// TIA Portal project "test_program" (V15)

(* hardware
DEVICE "S71500/ET200MP station_1"  S7-1500 station
   slot 0: "Rail_0"  Rack  6ES7 590-1***0-0AA0
   slot 0: "PM 70W 120/230VAC"  PM 70W 120/230VAC  6EP1332-4BA00
   slot 1: "PLC_1"  CPU 1511-1 PN  6ES7 511-1AK00-0AB0  V1.6
   slot 2: "DI 16x24VDC HF_1"  DI 16x24VDC HF  6ES7 521-1BH00-0AB0  V2.0
   slot 3: "DQ 16x24VDC/0.5A ST_1"  DQ 16x24VDC/0.5A ST  6ES7 522-1BH00-0AB0  V2.0
DEVICE "SCALANCE X005"  SCALANCE X-Station
   slot 0: "SCALANCE X rack"  Rail
   slot 0: "Switch_1"  6GK5 005-0BA00-1AA3  V1.0
DEVICE "GSD device_1"  GSD.Device.PN
   slot 0: "Rack"  Rack  V1.0
   slot 0: "INpactPIR"  Standard  INpact-PIR  V5.07
      slot 0: "Standard"  Standard
      slot 1: "Interface"  Interface
         slot 1: "Port 1"  Port 1
         slot 2: "Port 2"  Port 2
*)

// ===== PLC "PLC_1"  CPU 1511-1 PN =====
// protected blocks, not shown: "PDSql_1500_FB"

VAR_GLOBAL   // PLC tag table "Default tag table"
   "AlwaysTrue" AT %M0.1 : Bool;
   "AlwaysFalse" AT %M0.2 : Bool;
END_VAR

TYPE "part_processing_data"
   STRUCT
      sPartGroupID : String;
      rAFM_Param_1 : Real;
      rAFM_Param_2 : Real;
      rAFM_Param_3 : Real;
      sPartID_1 : String;
      iPartID_2 : UDInt;
   END_STRUCT;
END_TYPE

// folder: Data Types

TYPE "tConnection"
   STRUCT
      IP1 : USInt;
      IP2 : USInt;
      IP3 : USInt;
      IP4 : USInt;
      Port : UDInt;
      ConnID : Conn_Ouc;
      HW : Hw_Interface;
      Timeout : Time;
   END_STRUCT;
END_TYPE

TYPE "tSqlTable_1200"
   STRUCT
      ColumnCount : UInt;
      RowCount : UInt;
      MaxColumns : UInt := 10;
      MaxRows : UInt := 10;
      MaxStringLength : USInt := 50;
      Columns : Array[1..10] of "tColumn_1200";
   END_STRUCT;
END_TYPE

TYPE "tColumn_1200"
   STRUCT
      "Name" : String;   // Column name
      UserType : Byte;   // Unique generator of row
      "Type" : Byte;   // MSSQL-Data-Type of column
      LenSize : Byte;   // Number of bytes used for Length information of data
      TypeNumericPrecision : Byte;
      TypeNumericScale : Byte;
      Nullable : Bool;
      CaseSens : Bool;
      Identity : Bool;
      Computed : Bool;
      FixedLenCLRType : Bool;
      UsUpdatable : Byte;
      Rows : Array[1..10] of "tRow_1200";
   END_STRUCT;
END_TYPE

TYPE "tLicence"
   STRUCT
      LicKey1 : DWord;
      LicKey2 : DWord;
      LicKey3 : DWord;
      LicKey4 : DWord;
      LicKey5 : DWord;
   END_STRUCT;
END_TYPE

TYPE "tRow_1200"
   STRUCT
      "Bool" : Bool;
      Null : Bool;
      "DInt" : DInt;
      LReal : LReal;
      "String" : String[50];
      Datetime : DTL;
   END_STRUCT;
END_TYPE

TYPE "tSqlTable_1500"
   STRUCT
      ColumnCount : UInt;
      RowCount : UInt;
      MaxColumns : UInt := 10;
      MaxRows : UInt := 10;
      MaxStringLength : USInt := 50;
      Columns : Array[1..10] of "tColumn_1500";
   END_STRUCT;
END_TYPE

TYPE "tColumn_1500"
   STRUCT
      "Name" : String;   // Column name
      UserType : Byte;   // Unique generator of row
      "Type" : Byte;   // MSSQL-Data-Type of column
      LenSize : Byte;   // Number of bytes used for Length information of data
      TypeNumericPrecision : Byte;
      TypeNumericScale : Byte;
      Nullable : Bool;
      CaseSens : Bool;
      Identity : Bool;
      Computed : Bool;
      FixedLenCLRType : Bool;
      UsUpdatable : Byte;
      Rows : Array[1..10] of "tRow_1500";
   END_STRUCT;
END_TYPE

TYPE "tRow_1500"
   STRUCT
      "Bool" : Bool;
      Null : Bool;
      LInt : LInt;
      LReal : LReal;
      "String" : String[50];
      Datetime : DTL;
   END_STRUCT;
END_TYPE

TYPE "tLogin"
   STRUCT
      HostName : String[50];   // Hostname for database
      UserName : String[50];   // Username
      Password : String[50];   // Password
      Database : String[50];   // Database name
   END_STRUCT;
END_TYPE

TYPE "tQuery"
   STRUCT
      Query : Array[1..2] of String;
   END_STRUCT;
END_TYPE

TYPE "tCmd"
   STRUCT
      Connect : Bool;
      Disconnect : Bool;
      ExecuteQuery : Bool;
   END_STRUCT;
END_TYPE

TYPE "tStat"
   STRUCT
      Connected : Bool;
      Busy : Bool;
      ExecutedOK : Bool;
      Error : Bool;
      Status : Word;
      Message : String;
   END_STRUCT;
END_TYPE

// folder: 01_S7-1500

DATA_BLOCK "101_Simulation_IDB"   // DB1
{ S7_Optimized_Access := 'TRUE' }
VERSION : 0.1
// stored: InstanceOfName 101_Simulation
"101_Simulation"
BEGIN
END_DATA_BLOCK

DATA_BLOCK "InputsDB"   // DB2
{ S7_Optimized_Access := 'TRUE' }
VERSION : 0.1
   VAR
      part_processing_data : "part_processing_data";
   END_VAR
BEGIN
   part_processing_data.sPartGroupID := 'Deutz_ASML_10102A';
   part_processing_data.rAFM_Param_1 := 11.12;
   part_processing_data.rAFM_Param_2 := 4.98;
   part_processing_data.rAFM_Param_3 := 30.96;
   part_processing_data.sPartID_1 := 'ASML_JDK32_';
   part_processing_data.iPartID_2 := 100786;
END_DATA_BLOCK

DATA_BLOCK "DB_PDSql_1500"   // DB2010
{ S7_Optimized_Access := 'TRUE' }
VERSION : 0.1
   VAR
      Connection : "tConnection";
      Licence : "tLicence";
      Cmd : "tCmd";
      Stat : "tStat";
      Login : "tLogin";
      Query : "tQuery";
      SQLTable : "tSqlTable_1500";
   END_VAR
BEGIN
   Connection.IP1 := 192;
   Connection.IP2 := 168;
   Connection.IP3 := 2;
   Connection.IP4 := 1;
   Connection.Port := 1433;
   Login.Database := 'S7_1500_PLC';
   Login.Password := 'admin-6969';
   Login.UserName := 'sa';
   Login.HostName := 'EEEL1000332\SQLEXPRESS';
   Connection.ConnID := 1;
   Connection.HW := 64;
   Connection.Timeout := t#2s;
   Licence.LicKey1 := 16#67ABDCEB;
   Licence.LicKey2 := 16#28EC4AC9;
   Licence.LicKey3 := 16#D8D955FC;
   Licence.LicKey4 := 16#4A43863A;
   Licence.LicKey5 := 16#74F235FD;
END_DATA_BLOCK

// folder: 00_Functions

FUNCTION "LGF_Random_Real" : Real   // FC1, SCL
{ S7_Optimized_Access := 'TRUE' }
VERSION : 0.1
   VAR_OUTPUT
      error : Bool;
      status : Word;
      subfunctionStatus : Word;
   END_VAR
   VAR_TEMP
      tempTime : DTL;
      tempNanoSecondInDWord : DWord;
      tempTimeStatus : DWord;
      tempRandomValue : DWord;
   END_VAR
   VAR CONSTANT
      ZERO : Real;
      MAX_UDINT : UDInt := 4294967295;
      SUB_STATUS_NO_ERROR : Word := 16#0000;
      STATUS_FINISHED_NO_ERROR : Word := 16#0000;
      ERR_RD_SYS_T : Word := 16#8600;
   END_VAR
BEGIN
   REGION Block info header
       //=============================================================================
       // SIEMENS AG / (c)Copyright 2017
       //-----------------------------------------------------------------------------
       // Title:            LGF_Random_Real
       // Comment/Function: Generates a random real number between 0.0 and 1.0
       // Library/Family:   LGF(Library General Functions)
       // Author:           Siemens Digital Industry Support
       // Tested with:      S7-PLCSIM Advanced V2.0 SP1
       // Engineering:      TIA Portal V15 Update 2
       // Restrictions:     ENO disabled - error handling done by error and status
       // Requirements:     PLC (S7-1200 / S7-1500)
       //-------------------------------------------------------------------------------
       // Change log table:
       // Version  | Date       | Expert in charge       | Changes applied
       //----------|------------|------------------------|------------------------------
       // 01.00.00 27.01.2017  Siemens Industry Online Support
       //                      First released version
       // 01.00.01 17.08.2018  Siemens Industry Online Support
       //                      Upgrade: TIA V15 Update 2
       // 01.00.02 23.11.2018  Siemens Industry Online Support
       //                      Upgrade: TIA V15.1
       // 01.01.00 13.11.2019  Siemens Industry Presales Support
       //                      Renamed from "LGF_RandomBasic" to "LGF_Random_Real"
       //                      Regions, commens and costants are added
       // 03.00.00 23.04.2020  Siemens Industry Support
       //                      Set version to V3.0.0, harmonize the version of the whole library
       //=============================================================================
   END_REGION

   REGION Validation
       // Read system time
       #tempTimeStatus := INT_TO_WORD(RD_SYS_T(#tempTime));

       // Check return variable for error
       IF (#tempTimeStatus <> #SUB_STATUS_NO_ERROR) THEN
           #error := true;
           #status := #ERR_RD_SYS_T;
           #subfunctionStatus := #tempTimeStatus;
           #LGF_Random_Real := #ZERO;
           RETURN;
       END_IF;
   END_REGION

   REGION Calculating random number
       // Converting to double word so individual bytes can be addressed
       #tempNanoSecondInDWord := UDINT_TO_DWORD(#tempTime.NANOSECOND);

       // Calculate a random-start-value depending on the time
       #tempRandomValue.%B3 := #tempNanoSecondInDWord.%B0;
       #tempRandomValue.%B2 := #tempNanoSecondInDWord.%B1;
       #tempRandomValue.%B1 := #tempNanoSecondInDWord.%B2;
       #tempRandomValue.%B0 := #tempNanoSecondInDWord.%B3;

       // Norm the calculated random number: 0.0 <= Random_Real <= 1.0
       #LGF_Random_Real := UDINT_TO_REAL(DWORD_TO_UDINT(#tempRandomValue)) / UDINT_TO_REAL(#MAX_UDINT);

       #error := false;
       #status := #STATUS_FINISHED_NO_ERROR;
       #subfunctionStatus := #SUB_STATUS_NO_ERROR;
       // ENO mechanism is not used
       ENO := TRUE;
   END_REGION
END_FUNCTION

FUNCTION "fcRemovePlus" : String   // FC18, SCL
{ S7_Optimized_Access := 'TRUE' }
VERSION : 0.1
   VAR_INPUT
      STR : String;
   END_VAR
BEGIN
   //=============================================================================
   // PLCdirectSQL (c)Copyright 2019
   //-----------------------------------------------------------------------------
   // Library: fcRemovePlus
   // Tested with: S7-1200 FW 4.2 / S7-1500 FW 1.8
   // Engineering: TIA Portal 14
   // Requirements: S7-1200/1500
   // Functionality: Remove the first plus sign ("+") from a string
   //-----------------------------------------------------------------------------
   // Change log:
   // dd.mm.yyyy
   // 06.06.2019 Igor Filanda 1.0 First Release
   //=============================================================================

   IF FIND(IN1 := #STR, IN2 := '+') <> 0 THEN
       #fcRemovePlus := DELETE(IN := #STR, L := 1, P := FIND(IN1 := #STR, IN2 := '+'));
   ELSE
       #fcRemovePlus := #STR;
   END_IF;
END_FUNCTION

FUNCTION "fcDTLString" : String   // FC19, SCL
{ S7_Optimized_Access := 'TRUE' }
VERSION : 0.1
   VAR_INPUT
      dtlDatetime : DTL;
   END_VAR
   VAR_TEMP
      str : String;
   END_VAR
BEGIN
   //=============================================================================
   // PLCdirectSQL (c)Copyright 2019
   //-----------------------------------------------------------------------------
   // Library: fcDTLString
   // Tested with: S7-1200 FW 4.2 / S7-1500 FW 1.8
   // Engineering: TIA Portal 14
   // Requirements: S7-1200/1500
   // Functionality: Convert DTL data type (Datetime) to string
   //                (yyyy-MM-dd hh:mm:ss.fff)
   //-----------------------------------------------------------------------------
   // Change log:
   // dd.mm.yyyy
   // 06.06.2019 Igor Filanda 1.0 First Release
   //=============================================================================

   #str := "fcRemovePlus"(UDINT_TO_STRING(#dtlDatetime.YEAR));
   #str := CONCAT(IN1 := #str, IN2 := '-');
   #str := CONCAT(IN1 := #str, IN2 := "fcRemovePlus"(USINT_TO_STRING(#dtlDatetime.MONTH)));
   #str := CONCAT(IN1 := #str, IN2 := '-');
   #str := CONCAT(IN1 := #str, IN2 := "fcRemovePlus"(USINT_TO_STRING(#dtlDatetime.DAY)));
   #str := CONCAT(IN1 := #str, IN2 := ' ');
   #str := CONCAT(IN1 := #str, IN2 := "fcRemovePlus"(USINT_TO_STRING(#dtlDatetime.HOUR)));
   #str := CONCAT(IN1 := #str, IN2 := ':');
   #str := CONCAT(IN1 := #str, IN2 := "fcRemovePlus"(USINT_TO_STRING(#dtlDatetime.MINUTE)));
   #str := CONCAT(IN1 := #str, IN2 := ':');
   #str := CONCAT(IN1 := #str, IN2 := "fcRemovePlus"(USINT_TO_STRING(#dtlDatetime.SECOND)));
   #str := CONCAT(IN1 := #str, IN2 := '.');
   #str := CONCAT(IN1 := #str, IN2 := "fcRemovePlus"(UDINT_TO_STRING(#dtlDatetime.NANOSECOND / 1000000)));
   #fcDTLString := #str;
END_FUNCTION

// folder: 01_S7-1500

FUNCTION_BLOCK "101_Simulation"   // FB101, SCL
TITLE = 101_Simulation
{ S7_Optimized_Access := 'TRUE' }
VERSION : 0.1
   VAR
      State_101_Simulation : Int := 0;
      dtlDateTime : DTL;
      ton_1 : TON_TIME;
      ton_2 : TON_TIME;
      part_processing_data : "part_processing_data";
      bToggler : Bool;
      iToggler : Int;
   END_VAR
   VAR_TEMP
      "*************2" : Aom_Ident;
      sFruitName : String;
      iQuantity : Int;
      rWeight : Real;
      bCitrusType : Bool;
      "*************1" : Aom_Ident;
      str : String;
      LGF_Random_Real_error : Bool;
      LGF_Random_Real_status : Word;
      LGF_Random_Real_subfunctionStatus : Word;
      LGF_Random_Real : Real;
   END_VAR
BEGIN


   CASE #State_101_Simulation OF
       0:  //********************************
           #ton_1(IN:=TRUE,PT:=t#5000ms);
           IF #ton_1.Q THEN
               #ton_1(IN := FALSE,PT := t#0s);
               #State_101_Simulation := 10;
           END_IF;

       10: //********************************
           #LGF_Random_Real:= "LGF_Random_Real"(error=>#LGF_Random_Real_error,
                                                status=>#LGF_Random_Real_status,
                                                subfunctionStatus=>#LGF_Random_Real_subfunctionStatus);
           #bToggler := NOT #bToggler;
           IF #bToggler = TRUE THEN
               #iToggler := 1;
           ELSE
               #iToggler := -1;
           END_IF;

           //*********************************
           #part_processing_data.sPartGroupID := "InputsDB".part_processing_data.sPartGroupID;
           #part_processing_data.rAFM_Param_1 := "InputsDB".#part_processing_data.rAFM_Param_1+ (#LGF_Random_Real*#iToggler);
           #part_processing_data.rAFM_Param_2 := "InputsDB".part_processing_data.#rAFM_Param_2+ (#LGF_Random_Real*#iToggler);
           #part_processing_data.rAFM_Param_3 := "InputsDB".part_processing_data.#rAFM_Param_3+ (#LGF_Random_Real*#iToggler);
           "InputsDB".part_processing_data.iPartID_2 := "InputsDB".part_processing_data.iPartID_2+1;
           #part_processing_data.sPartID_1 := CONCAT(IN1 := "InputsDB".part_processing_data.sPartID_1,
                                                     IN2 := "fcRemovePlus"(UDINT_TO_STRING("InputsDB".part_processing_data.iPartID_2)));

           // DO NOT FORGET TO UPDATE YOUR [TABLE NAME](e.g. TestTable1) IN THE BELOW FIRST STRING !
           #str := 'INSERT INTO TestTable1(Datetime,PartGroupID,AFM_Param_1,AFM_Param_2,AFM_Param_3,PartID) VALUES($'';
           #str := CONCAT(IN1 := #str, IN2 := "fcDTLString"(#dtlDateTime));
           #str := CONCAT(IN1 := #str, IN2 := '$',$'');
           #str := CONCAT(IN1 := #str, IN2 := #part_processing_data.sPartGroupID);
           #str := CONCAT(IN1 := #str, IN2 := '$',');
           #str := CONCAT(IN1 := #str, IN2 := REAL_TO_STRING(#part_processing_data.rAFM_Param_1));
           #str := CONCAT(IN1 := #str, IN2 := ',');
           #str := CONCAT(IN1 := #str, IN2 := REAL_TO_STRING(#part_processing_data.rAFM_Param_2));
           #str := CONCAT(IN1 := #str, IN2 := ',');
           #str := CONCAT(IN1 := #str, IN2 := REAL_TO_STRING(#part_processing_data.rAFM_Param_3));
           #str := CONCAT(IN1 := #str, IN2 := ',');
           #str := CONCAT(IN1 := #str, IN2 := '$'');
           #str := CONCAT(IN1 := #str, IN2 := #part_processing_data.sPartID_1);
           #str := CONCAT(IN1 := #str, IN2 := '$'');
           #str := CONCAT(IN1 := #str, IN2 := ')');

           "DB_PDSql_1500".Query.Query[1] := #str;
           "DB_PDSql_1500".Query.Query[2] := '';
           IF TRUE THEN
               "DB_PDSql_1500".Cmd.ExecuteQuery := TRUE;
               #State_101_Simulation := 100;
           END_IF;

       100:  //********************************
           #ton_1(IN := TRUE,PT := t#5000ms);
           IF #ton_1.Q AND TRUE THEN
               #ton_1(IN := FALSE,PT := t#0s);
               "DB_PDSql_1500".Cmd.ExecuteQuery := FALSE;
               #State_101_Simulation := 0;
           END_IF;


       ELSE  // Statement section ELSE
           ;
   END_CASE;
END_FUNCTION_BLOCK

ORGANIZATION_BLOCK "Main"   // OB1, LAD, ProgramCycle
TITLE = "Main Program Sweep (Cycle)"
{ S7_Optimized_Access := 'TRUE' }
VERSION : 0.1
   VAR_INPUT
      Initial_Call : Bool;   // Initial call of this OB
      Remanence : Bool;   // =True, if remanent data are available
   END_VAR
   VAR_TEMP
      RetVal : Word;
      OUT : DTL;
   END_VAR
BEGIN

REGION Network 1: PDSql Library
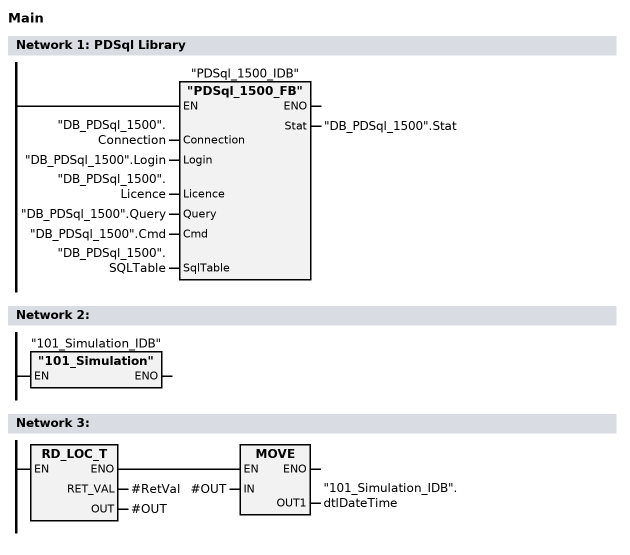
   RUNG wire#powerrail
      "PDSql_1500_IDB"(Connection := "DB_PDSql_1500".Connection, Login := "DB_PDSql_1500".Login, Licence := "DB_PDSql_1500".Licence, Query := "DB_PDSql_1500".Query, Cmd := "DB_PDSql_1500".Cmd, SqlTable := "DB_PDSql_1500".SQLTable, Stat => "DB_PDSql_1500".Stat)
   END_RUNG
   // the same network as SCL:
   "PDSql_1500_IDB"(Connection := "DB_PDSql_1500".Connection,   // "PDSql_1500_FB"
                    Login := "DB_PDSql_1500".Login,
                    Licence := "DB_PDSql_1500".Licence,
                    Query := "DB_PDSql_1500".Query,
                    Cmd := "DB_PDSql_1500".Cmd,
                    SqlTable := "DB_PDSql_1500".SQLTable,
                    Stat => "DB_PDSql_1500".Stat);
END_REGION

REGION Network 2
   RUNG wire#powerrail
      "101_Simulation_IDB"()
   END_RUNG
   // the same network as SCL:
   "101_Simulation_IDB"();   // "101_Simulation"
END_REGION

REGION Network 3
   // ENO of a box is taken as its EN; it also drops when the box reports an error
   #RetVal := RD_LOC_T(OUT => #OUT);
   "101_Simulation_IDB".dtlDateTime := #OUT;
END_REGION
END_ORGANIZATION_BLOCK

// ===== library: CodeBlockByCopyVersionObject "None" =====
// protected blocks, not shown: "hg1jahs3gd0jgsa1ba671de-d280-4bff-a15f-7f20c6828afd0"

// ===== library: CodeBlockByCopyVersionObject "None" =====
// protected blocks, not shown: "hg1jahs3gd0jgsa9326f056-fdd1-4983-8b45-f083db44157f0"